   2973: 'Carrier 46 Power unit: Line phase failure in main circuit', class No Acknowledgement, trigger "DB302_HMI_Faults_Carrier46_Faults_1" bit 12
   2974: 'Carrier 46 Power unit: Phase failure motor cable', class No Acknowledgement, trigger "DB302_HMI_Faults_Carrier46_Faults_1" bit 13
   2975: 'Carrier 46 Power unit: Ground fault', class No Acknowledgement, trigger "DB302_HMI_Faults_Carrier46_Faults_1" bit 14
   2976: 'Spare_Fault_2976', class No Acknowledgement, trigger "DB302_HMI_Faults_Carrier46_Faults_1" bit 15
   2977: 'Carrier 46 Motion Off Fault', class No Acknowledgement, trigger "DB302_HMI_Faults_Carrier46_Faults_2" bit 0
   2978: 'Carrier 46 Motion On Fault', class No Acknowledgement, trigger "DB302_HMI_Faults_Carrier46_Faults_2" bit 1
   2979: 'Carrier 46 Spacing Fault', class No Acknowledgement, trigger "DB302_HMI_Faults_Carrier46_Faults_2" bit 2
   2980: 'Carrier 46 Duplicate Carrier Number Fault', class No Acknowledgement, trigger "DB302_HMI_Faults_Carrier46_Faults_2" bit 3
   2981: 'Spare_Fault_2981', class No Acknowledgement, trigger "DB302_HMI_Faults_Carrier46_Faults_2" bit 4
   2982: 'Spare_Fault_2982', class No Acknowledgement, trigger "DB302_HMI_Faults_Carrier46_Faults_2" bit 5
   2983: 'Spare_Fault_2983', class No Acknowledgement, trigger "DB302_HMI_Faults_Carrier46_Faults_2" bit 6
   2984: 'Spare_Fault_2984', class No Acknowledgement, trigger "DB302_HMI_Faults_Carrier46_Faults_2" bit 7
   2985: 'Spare_Fault_2985', class No Acknowledgement, trigger "DB302_HMI_Faults_Carrier46_Faults_2" bit 8
   2986: 'Spare_Fault_2986', class No Acknowledgement, trigger "DB302_HMI_Faults_Carrier46_Faults_2" bit 9
   2987: 'Spare_Fault_2987', class No Acknowledgement, trigger "DB302_HMI_Faults_Carrier46_Faults_2" bit 10
   2988: 'Spare_Fault_2988', class No Acknowledgement, trigger "DB302_HMI_Faults_Carrier46_Faults_2" bit 11
   2989: 'Spare_Fault_2989', class No Acknowledgement, trigger "DB302_HMI_Faults_Carrier46_Faults_2" bit 12
   2990: 'Spare_Fault_2990', class No Acknowledgement, trigger "DB302_HMI_Faults_Carrier46_Faults_2" bit 13
   2991: 'Spare_Fault_2991', class No Acknowledgement, trigger "DB302_HMI_Faults_Carrier46_Faults_2" bit 14
   2992: 'Spare_Fault_2992', class No Acknowledgement, trigger "DB302_HMI_Faults_Carrier46_Faults_2" bit 15
   2993: 'Spare_Fault_2993', class No Acknowledgement, trigger "DB302_HMI_Faults_Carrier46_Faults_3" bit 0
   2994: 'Spare_Fault_2994', class No Acknowledgement, trigger "DB302_HMI_Faults_Carrier46_Faults_3" bit 1
   2995: 'Spare_Fault_2995', class No Acknowledgement, trigger "DB302_HMI_Faults_Carrier46_Faults_3" bit 2
   2996: 'Spare_Fault_2996', class No Acknowledgement, trigger "DB302_HMI_Faults_Carrier46_Faults_3" bit 3
   2997: 'Spare_Fault_2997', class No Acknowledgement, trigger "DB302_HMI_Faults_Carrier46_Faults_3" bit 4
   2998: 'Spare_Fault_2998', class No Acknowledgement, trigger "DB302_HMI_Faults_Carrier46_Faults_3" bit 5
   2999: 'Spare_Fault_2999', class No Acknowledgement, trigger "DB302_HMI_Faults_Carrier46_Faults_3" bit 6
   3000: 'Spare_Fault_3000', class No Acknowledgement, trigger "DB302_HMI_Faults_Carrier46_Faults_3" bit 7
   3001: 'Spare_Fault_3001', class No Acknowledgement, trigger "DB302_HMI_Faults_Carrier46_Faults_3" bit 8
   3002: 'Spare_Fault_3002', class No Acknowledgement, trigger "DB302_HMI_Faults_Carrier46_Faults_3" bit 9
   3003: 'Spare_Fault_3003', class No Acknowledgement, trigger "DB302_HMI_Faults_Carrier46_Faults_3" bit 10
   3004: 'Spare_Fault_3004', class No Acknowledgement, trigger "DB302_HMI_Faults_Carrier46_Faults_3" bit 11
   3005: 'Spare_Fault_3005', class No Acknowledgement, trigger "DB302_HMI_Faults_Carrier46_Faults_3" bit 12
   3006: 'Spare_Fault_3006', class No Acknowledgement, trigger "DB302_HMI_Faults_Carrier46_Faults_3" bit 13
   3007: 'Spare_Fault_3007', class No Acknowledgement, trigger "DB302_HMI_Faults_Carrier46_Faults_3" bit 14
   3008: 'Spare_Fault_3008', class No Acknowledgement, trigger "DB302_HMI_Faults_Carrier46_Faults_3" bit 15
   3009: 'Carrier 47 Disconnect Open Power Fault DI11.0', class No Acknowledgement, trigger "DB302_HMI_Faults_Carrier47_Faults_0" bit 0
   3010: 'Carrier 47 Drive Profinet Comm Fault', class No Acknowledgement, trigger "DB302_HMI_Faults_Carrier47_Faults_0" bit 1
   3011: 'Carrier 47 Production Stop Not Reset', class No Acknowledgement, trigger "DB302_HMI_Faults_Carrier47_Faults_0" bit 2
   3012: 'Carrier 47 CB02122 Tripped', class No Acknowledgement, trigger "DB302_HMI_Faults_Carrier47_Faults_0" bit 3
   3013: 'Carrier 47 CB02123 Tripped', class No Acknowledgement, trigger "DB302_HMI_Faults_Carrier47_Faults_0" bit 4
   3014: 'Carrier 47 AUX1 CB Tripped', class No Acknowledgement, trigger "DB302_HMI_Faults_Carrier47_Faults_0" bit 5
   3015: 'Carrier 47 AUX2 CB Tripped', class No Acknowledgement, trigger "DB302_HMI_Faults_Carrier47_Faults_0" bit 6
   3016: 'Carrier 47 PLC Not Communicating', class No Acknowledgement, trigger "DB302_HMI_Faults_Carrier47_Faults_0" bit 7
   3017: 'Carrier 47 Safe Input Card Fault', class No Acknowledgement, trigger "DB302_HMI_Faults_Carrier47_Faults_0" bit 8
   3018: 'Carrier 47 Safe Output Card Fault', class No Acknowledgement, trigger "DB302_HMI_Faults_Carrier47_Faults_0" bit 9
   3019: 'Carrier 47 Standard Input Card Fault', class No Acknowledgement, trigger "DB302_HMI_Faults_Carrier47_Faults_0" bit 10
   3020: 'Carrier 47 Standard Output Card Fault', class No Acknowledgement, trigger "DB302_HMI_Faults_Carrier47_Faults_0" bit 11
   3021: 'Carrier 47 Encoder Position Fault', class No Acknowledgement, trigger "DB302_HMI_Faults_Carrier47_Faults_0" bit 12
   3022: 'Carrier 47 Encoder Internal Error', class No Acknowledgement, trigger "DB302_HMI_Faults_Carrier47_Faults_0" bit 13
   3023: 'Carrier 47 Encoder Comm Fault', class No Acknowledgement, trigger "DB302_HMI_Faults_Carrier47_Faults_0" bit 14
   3024: 'Carrier 47 HMI Comm Fault', class No Acknowledgement, trigger "DB302_HMI_Faults_Carrier47_Faults_0" bit 15
   3025: 'Carrier 47 Crash Detection Fault', class No Acknowledgement, trigger "DB302_HMI_Faults_Carrier47_Faults_1" bit 0
   3026: 'Carrier 47 Carrier Number Invalid', class No Acknowledgement, trigger "DB302_HMI_Faults_Carrier47_Faults_1" bit 1
   3027: 'Carrier 47 Drive: PROFINET configuration error', class No Acknowledgement, trigger "DB302_HMI_Faults_Carrier47_Faults_1" bit 2
   3028: 'Carrier 47 Drive: Error internal communications', class No Acknowledgement, trigger "DB302_HMI_Faults_Carrier47_Faults_1" bit 3
   3029: 'Carrier 47 Drive: Motor overtemperature', class No Acknowledgement, trigger "DB302_HMI_Faults_Carrier47_Faults_1" bit 4
   3030: 'Carrier 47 Drive: Motor overcurrent', class No Acknowledgement, trigger "DB302_HMI_Faults_Carrier47_Faults_1" bit 5
   3031: 'Carrier 47 Drive: Infeed or power unit not ready', class No Acknowledgement, trigger "DB302_HMI_Faults_Carrier47_Faults_1" bit 6
   3032: 'Carrier 47 Drive: Short-circuit/ground fault detected', class No Acknowledgement, trigger "DB302_HMI_Faults_Carrier47_Faults_1" bit 7
   3033: 'Carrier 47 Drive: PROFINET Setpoint timeout', class No Acknowledgement, trigger "DB302_HMI_Faults_Carrier47_Faults_1" bit 8
   3034: 'Carrier 47 Power unit: Overcurrent', class No Acknowledgement, trigger "DB302_HMI_Faults_Carrier47_Faults_1" bit 9
   3035: 'Carrier 47 Power unit: DC link voltage overvoltage', class No Acknowledgement, trigger "DB302_HMI_Faults_Carrier47_Faults_1" bit 10
   3036: 'Carrier 47 Power unit: DC link voltage undervoltage', class No Acknowledgement, trigger "DB302_HMI_Faults_Carrier47_Faults_1" bit 11
   3037: 'Carrier 47 Power unit: Line phase failure in main circuit', class No Acknowledgement, trigger "DB302_HMI_Faults_Carrier47_Faults_1" bit 12
   3038: 'Carrier 47 Power unit: Phase failure motor cable', class No Acknowledgement, trigger "DB302_HMI_Faults_Carrier47_Faults_1" bit 13
   3039: 'Carrier 47 Power unit: Ground fault', class No Acknowledgement, trigger "DB302_HMI_Faults_Carrier47_Faults_1" bit 14
   3040: 'Spare_Fault_3040', class No Acknowledgement, trigger "DB302_HMI_Faults_Carrier47_Faults_1" bit 15
   3041: 'Carrier 47 Motion Off Fault', class No Acknowledgement, trigger "DB302_HMI_Faults_Carrier47_Faults_2" bit 0
   3042: 'Carrier 47 Motion On Fault', class No Acknowledgement, trigger "DB302_HMI_Faults_Carrier47_Faults_2" bit 1
   3043: 'Carrier 47 Spacing Fault', class No Acknowledgement, trigger "DB302_HMI_Faults_Carrier47_Faults_2" bit 2
   3044: 'Carrier 47 Duplicate Carrier Number Fault', class No Acknowledgement, trigger "DB302_HMI_Faults_Carrier47_Faults_2" bit 3
   3045: 'Spare_Fault_3045', class No Acknowledgement, trigger "DB302_HMI_Faults_Carrier47_Faults_2" bit 4
   3046: 'Spare_Fault_3046', class No Acknowledgement, trigger "DB302_HMI_Faults_Carrier47_Faults_2" bit 5
   3047: 'Spare_Fault_3047', class No Acknowledgement, trigger "DB302_HMI_Faults_Carrier47_Faults_2" bit 6
   3048: 'Spare_Fault_3048', class No Acknowledgement, trigger "DB302_HMI_Faults_Carrier47_Faults_2" bit 7
   3049: 'Spare_Fault_3049', class No Acknowledgement, trigger "DB302_HMI_Faults_Carrier47_Faults_2" bit 8
   3050: 'Spare_Fault_3050', class No Acknowledgement, trigger "DB302_HMI_Faults_Carrier47_Faults_2" bit 9
   3051: 'Spare_Fault_3051', class No Acknowledgement, trigger "DB302_HMI_Faults_Carrier47_Faults_2" bit 10
   3052: 'Spare_Fault_3052', class No Acknowledgement, trigger "DB302_HMI_Faults_Carrier47_Faults_2" bit 11
   3053: 'Spare_Fault_3053', class No Acknowledgement, trigger "DB302_HMI_Faults_Carrier47_Faults_2" bit 12
   3054: 'Spare_Fault_3054', class No Acknowledgement, trigger "DB302_HMI_Faults_Carrier47_Faults_2" bit 13
   3055: 'Spare_Fault_3055', class No Acknowledgement, trigger "DB302_HMI_Faults_Carrier47_Faults_2" bit 14
   3056: 'Spare_Fault_3056', class No Acknowledgement, trigger "DB302_HMI_Faults_Carrier47_Faults_2" bit 15
   3057: 'Spare_Fault_3057', class No Acknowledgement, trigger "DB302_HMI_Faults_Carrier47_Faults_3" bit 0
   3058: 'Spare_Fault_3058', class No Acknowledgement, trigger "DB302_HMI_Faults_Carrier47_Faults_3" bit 1
   3059: 'Spare_Fault_3059', class No Acknowledgement, trigger "DB302_HMI_Faults_Carrier47_Faults_3" bit 2
   3060: 'Spare_Fault_3060', class No Acknowledgement, trigger "DB302_HMI_Faults_Carrier47_Faults_3" bit 3
   3061: 'Spare_Fault_3061', class No Acknowledgement, trigger "DB302_HMI_Faults_Carrier47_Faults_3" bit 4
   3062: 'Spare_Fault_3062', class No Acknowledgement, trigger "DB302_HMI_Faults_Carrier47_Faults_3" bit 5
   3063: 'Spare_Fault_3063', class No Acknowledgement, trigger "DB302_HMI_Faults_Carrier47_Faults_3" bit 6
   3064: 'Spare_Fault_3064', class No Acknowledgement, trigger "DB302_HMI_Faults_Carrier47_Faults_3" bit 7
   3065: 'Spare_Fault_3065', class No Acknowledgement, trigger "DB302_HMI_Faults_Carrier47_Faults_3" bit 8
   3066: 'Spare_Fault_3066', class No Acknowledgement, trigger "DB302_HMI_Faults_Carrier47_Faults_3" bit 9
   3067: 'Spare_Fault_3067', class No Acknowledgement, trigger "DB302_HMI_Faults_Carrier47_Faults_3" bit 10
   3068: 'Spare_Fault_3068', class No Acknowledgement, trigger "DB302_HMI_Faults_Carrier47_Faults_3" bit 11
   3069: 'Spare_Fault_3069', class No Acknowledgement, trigger "DB302_HMI_Faults_Carrier47_Faults_3" bit 12
   3070: 'Spare_Fault_3070', class No Acknowledgement, trigger "DB302_HMI_Faults_Carrier47_Faults_3" bit 13
   3071: 'Spare_Fault_3071', class No Acknowledgement, trigger "DB302_HMI_Faults_Carrier47_Faults_3" bit 14
   3072: 'Spare_Fault_3072', class No Acknowledgement, trigger "DB302_HMI_Faults_Carrier47_Faults_3" bit 15
   3073: 'Carrier 48 Disconnect Open Power Fault DI11.0', class No Acknowledgement, trigger "DB302_HMI_Faults_Carrier48_Faults_0" bit 0
   3074: 'Carrier 48 Drive Profinet Comm Fault', class No Acknowledgement, trigger "DB302_HMI_Faults_Carrier48_Faults_0" bit 1
   3075: 'Carrier 48 Production Stop Not Reset', class No Acknowledgement, trigger "DB302_HMI_Faults_Carrier48_Faults_0" bit 2
   3076: 'Carrier 48 CB02122 Tripped', class No Acknowledgement, trigger "DB302_HMI_Faults_Carrier48_Faults_0" bit 3
   3077: 'Carrier 48 CB02123 Tripped', class No Acknowledgement, trigger "DB302_HMI_Faults_Carrier48_Faults_0" bit 4
   3078: 'Carrier 48 AUX1 CB Tripped', class No Acknowledgement, trigger "DB302_HMI_Faults_Carrier48_Faults_0" bit 5
   3079: 'Carrier 48 AUX2 CB Tripped', class No Acknowledgement, trigger "DB302_HMI_Faults_Carrier48_Faults_0" bit 6
   3080: 'Carrier 48 PLC Not Communicating', class No Acknowledgement, trigger "DB302_HMI_Faults_Carrier48_Faults_0" bit 7
   3081: 'Carrier 48 Safe Input Card Fault', class No Acknowledgement, trigger "DB302_HMI_Faults_Carrier48_Faults_0" bit 8
   3082: 'Carrier 48 Safe Output Card Fault', class No Acknowledgement, trigger "DB302_HMI_Faults_Carrier48_Faults_0" bit 9
   3083: 'Carrier 48 Standard Input Card Fault', class No Acknowledgement, trigger "DB302_HMI_Faults_Carrier48_Faults_0" bit 10
   3084: 'Carrier 48 Standard Output Card Fault', class No Acknowledgement, trigger "DB302_HMI_Faults_Carrier48_Faults_0" bit 11
   3085: 'Carrier 48 Encoder Position Fault', class No Acknowledgement, trigger "DB302_HMI_Faults_Carrier48_Faults_0" bit 12
   3086: 'Carrier 48 Encoder Internal Error', class No Acknowledgement, trigger "DB302_HMI_Faults_Carrier48_Faults_0" bit 13
   3087: 'Carrier 48 Encoder Comm Fault', class No Acknowledgement, trigger "DB302_HMI_Faults_Carrier48_Faults_0" bit 14
   3088: 'Carrier 48 HMI Comm Fault', class No Acknowledgement, trigger "DB302_HMI_Faults_Carrier48_Faults_0" bit 15
   3089: 'Carrier 48 Crash Detection Fault', class No Acknowledgement, trigger "DB302_HMI_Faults_Carrier48_Faults_1" bit 0
   3090: 'Carrier 48 Carrier Number Invalid', class No Acknowledgement, trigger "DB302_HMI_Faults_Carrier48_Faults_1" bit 1
   3091: 'Carrier 48 Drive: PROFINET configuration error', class No Acknowledgement, trigger "DB302_HMI_Faults_Carrier48_Faults_1" bit 2
   3092: 'Carrier 48 Drive: Error internal communications', class No Acknowledgement, trigger "DB302_HMI_Faults_Carrier48_Faults_1" bit 3
   3093: 'Carrier 48 Drive: Motor overtemperature', class No Acknowledgement, trigger "DB302_HMI_Faults_Carrier48_Faults_1" bit 4
   3094: 'Carrier 48 Drive: Motor overcurrent', class No Acknowledgement, trigger "DB302_HMI_Faults_Carrier48_Faults_1" bit 5
   3095: 'Carrier 48 Drive: Infeed or power unit not ready', class No Acknowledgement, trigger "DB302_HMI_Faults_Carrier48_Faults_1" bit 6
   3096: 'Carrier 48 Drive: Short-circuit/ground fault detected', class No Acknowledgement, trigger "DB302_HMI_Faults_Carrier48_Faults_1" bit 7
   3097: 'Carrier 48 Drive: PROFINET Setpoint timeout', class No Acknowledgement, trigger "DB302_HMI_Faults_Carrier48_Faults_1" bit 8
   3098: 'Carrier 48 Power unit: Overcurrent', class No Acknowledgement, trigger "DB302_HMI_Faults_Carrier48_Faults_1" bit 9
   3099: 'Carrier 48 Power unit: DC link voltage overvoltage', class No Acknowledgement, trigger "DB302_HMI_Faults_Carrier48_Faults_1" bit 10
   3100: 'Carrier 48 Power unit: DC link voltage undervoltage', class No Acknowledgement, trigger "DB302_HMI_Faults_Carrier48_Faults_1" bit 11
   3101: 'Carrier 48 Power unit: Line phase failure in main circuit', class No Acknowledgement, trigger "DB302_HMI_Faults_Carrier48_Faults_1" bit 12
   3102: 'Carrier 48 Power unit: Phase failure motor cable', class No Acknowledgement, trigger "DB302_HMI_Faults_Carrier48_Faults_1" bit 13
   3103: 'Carrier 48 Power unit: Ground fault', class No Acknowledgement, trigger "DB302_HMI_Faults_Carrier48_Faults_1" bit 14
   3104: 'Spare_Fault_3104', class No Acknowledgement, trigger "DB302_HMI_Faults_Carrier48_Faults_1" bit 15
   3105: 'Carrier 48 Motion Off Fault', class No Acknowledgement, trigger "DB302_HMI_Faults_Carrier48_Faults_2" bit 0
   3106: 'Carrier 48 Motion On Fault', class No Acknowledgement, trigger "DB302_HMI_Faults_Carrier48_Faults_2" bit 1
   3107: 'Carrier 48 Spacing Fault', class No Acknowledgement, trigger "DB302_HMI_Faults_Carrier48_Faults_2" bit 2
   3108: 'Carrier 48 Duplicate Carrier Number Fault', class No Acknowledgement, trigger "DB302_HMI_Faults_Carrier48_Faults_2" bit 3
   3109: 'Spare_Fault_3109', class No Acknowledgement, trigger "DB302_HMI_Faults_Carrier48_Faults_2" bit 4
   3110: 'Spare_Fault_3110', class No Acknowledgement, trigger "DB302_HMI_Faults_Carrier48_Faults_2" bit 5
   3111: 'Spare_Fault_3111', class No Acknowledgement, trigger "DB302_HMI_Faults_Carrier48_Faults_2" bit 6
   3112: 'Spare_Fault_3112', class No Acknowledgement, trigger "DB302_HMI_Faults_Carrier48_Faults_2" bit 7
   3113: 'Spare_Fault_3113', class No Acknowledgement, trigger "DB302_HMI_Faults_Carrier48_Faults_2" bit 8
   3114: 'Spare_Fault_3114', class No Acknowledgement, trigger "DB302_HMI_Faults_Carrier48_Faults_2" bit 9
   3115: 'Spare_Fault_3115', class No Acknowledgement, trigger "DB302_HMI_Faults_Carrier48_Faults_2" bit 10
   3116: 'Spare_Fault_3116', class No Acknowledgement, trigger "DB302_HMI_Faults_Carrier48_Faults_2" bit 11
   3117: 'Spare_Fault_3117', class No Acknowledgement, trigger "DB302_HMI_Faults_Carrier48_Faults_2" bit 12
   3118: 'Spare_Fault_3118', class No Acknowledgement, trigger "DB302_HMI_Faults_Carrier48_Faults_2" bit 13
   3119: 'Spare_Fault_3119', class No Acknowledgement, trigger "DB302_HMI_Faults_Carrier48_Faults_2" bit 14
   3120: 'Spare_Fault_3120', class No Acknowledgement, trigger "DB302_HMI_Faults_Carrier48_Faults_2" bit 15
   3121: 'Spare_Fault_3121', class No Acknowledgement, trigger "DB302_HMI_Faults_Carrier48_Faults_3" bit 0
   3122: 'Spare_Fault_3122', class No Acknowledgement, trigger "DB302_HMI_Faults_Carrier48_Faults_3" bit 1
   3123: 'Spare_Fault_3123', class No Acknowledgement, trigger "DB302_HMI_Faults_Carrier48_Faults_3" bit 2
   3124: 'Spare_Fault_3124', class No Acknowledgement, trigger "DB302_HMI_Faults_Carrier48_Faults_3" bit 3
   3125: 'Spare_Fault_3125', class No Acknowledgement, trigger "DB302_HMI_Faults_Carrier48_Faults_3" bit 4
   3126: 'Spare_Fault_3126', class No Acknowledgement, trigger "DB302_HMI_Faults_Carrier48_Faults_3" bit 5
   3127: 'Spare_Fault_3127', class No Acknowledgement, trigger "DB302_HMI_Faults_Carrier48_Faults_3" bit 6
   3128: 'Spare_Fault_3128', class No Acknowledgement, trigger "DB302_HMI_Faults_Carrier48_Faults_3" bit 7
   3129: 'Spare_Fault_3129', class No Acknowledgement, trigger "DB302_HMI_Faults_Carrier48_Faults_3" bit 8
   3130: 'Spare_Fault_3130', class No Acknowledgement, trigger "DB302_HMI_Faults_Carrier48_Faults_3" bit 9
   3131: 'Spare_Fault_3131', class No Acknowledgement, trigger "DB302_HMI_Faults_Carrier48_Faults_3" bit 10
   3132: 'Spare_Fault_3132', class No Acknowledgement, trigger "DB302_HMI_Faults_Carrier48_Faults_3" bit 11
   3133: 'Spare_Fault_3133', class No Acknowledgement, trigger "DB302_HMI_Faults_Carrier48_Faults_3" bit 12
   3134: 'Spare_Fault_3134', class No Acknowledgement, trigger "DB302_HMI_Faults_Carrier48_Faults_3" bit 13
   3135: 'Spare_Fault_3135', class No Acknowledgement, trigger "DB302_HMI_Faults_Carrier48_Faults_3" bit 14
   3136: 'Spare_Fault_3136', class No Acknowledgement, trigger "DB302_HMI_Faults_Carrier48_Faults_3" bit 15
   3137: 'Carrier 49 Disconnect Open Power Fault DI11.0', class No Acknowledgement, trigger "DB302_HMI_Faults_Carrier49_Faults_0" bit 0
   3138: 'Carrier 49 Drive Profinet Comm Fault', class No Acknowledgement, trigger "DB302_HMI_Faults_Carrier49_Faults_0" bit 1
   3139: 'Carrier 49 Production Stop Not Reset', class No Acknowledgement, trigger "DB302_HMI_Faults_Carrier49_Faults_0" bit 2
   3140: 'Carrier 49 CB02122 Tripped', class No Acknowledgement, trigger "DB302_HMI_Faults_Carrier49_Faults_0" bit 3
   3141: 'Carrier 49 CB02123 Tripped', class No Acknowledgement, trigger "DB302_HMI_Faults_Carrier49_Faults_0" bit 4
   3142: 'Carrier 49 AUX1 CB Tripped', class No Acknowledgement, trigger "DB302_HMI_Faults_Carrier49_Faults_0" bit 5
   3143: 'Carrier 49 AUX2 CB Tripped', class No Acknowledgement, trigger "DB302_HMI_Faults_Carrier49_Faults_0" bit 6
   3144: 'Carrier 49 PLC Not Communicating', class No Acknowledgement, trigger "DB302_HMI_Faults_Carrier49_Faults_0" bit 7
   3145: 'Carrier 49 Safe Input Card Fault', class No Acknowledgement, trigger "DB302_HMI_Faults_Carrier49_Faults_0" bit 8
   3146: 'Carrier 49 Safe Output Card Fault', class No Acknowledgement, trigger "DB302_HMI_Faults_Carrier49_Faults_0" bit 9
   3147: 'Carrier 49 Standard Input Card Fault', class No Acknowledgement, trigger "DB302_HMI_Faults_Carrier49_Faults_0" bit 10
   3148: 'Carrier 49 Standard Output Card Fault', class No Acknowledgement, trigger "DB302_HMI_Faults_Carrier49_Faults_0" bit 11
   3149: 'Carrier 49 Encoder Position Fault', class No Acknowledgement, trigger "DB302_HMI_Faults_Carrier49_Faults_0" bit 12
   3150: 'Carrier 49 Encoder Internal Error', class No Acknowledgement, trigger "DB302_HMI_Faults_Carrier49_Faults_0" bit 13
   3151: 'Carrier 49 Encoder Comm Fault', class No Acknowledgement, trigger "DB302_HMI_Faults_Carrier49_Faults_0" bit 14
   3152: 'Carrier 49 HMI Comm Fault', class No Acknowledgement, trigger "DB302_HMI_Faults_Carrier49_Faults_0" bit 15
   3153: 'Carrier 49 Crash Detection Fault', class No Acknowledgement, trigger "DB302_HMI_Faults_Carrier49_Faults_1" bit 0
   3154: 'Carrier 49 Carrier Number Invalid', class No Acknowledgement, trigger "DB302_HMI_Faults_Carrier49_Faults_1" bit 1
   3155: 'Carrier 49 Drive: PROFINET configuration error', class No Acknowledgement, trigger "DB302_HMI_Faults_Carrier49_Faults_1" bit 2
   3156: 'Carrier 49 Drive: Error internal communications', class No Acknowledgement, trigger "DB302_HMI_Faults_Carrier49_Faults_1" bit 3
   3157: 'Carrier 49 Drive: Motor overtemperature', class No Acknowledgement, trigger "DB302_HMI_Faults_Carrier49_Faults_1" bit 4
   3158: 'Carrier 49 Drive: Motor overcurrent', class No Acknowledgement, trigger "DB302_HMI_Faults_Carrier49_Faults_1" bit 5
   3159: 'Carrier 49 Drive: Infeed or power unit not ready', class No Acknowledgement, trigger "DB302_HMI_Faults_Carrier49_Faults_1" bit 6
   3160: 'Carrier 49 Drive: Short-circuit/ground fault detected', class No Acknowledgement, trigger "DB302_HMI_Faults_Carrier49_Faults_1" bit 7
   3161: 'Carrier 49 Drive: PROFINET Setpoint timeout', class No Acknowledgement, trigger "DB302_HMI_Faults_Carrier49_Faults_1" bit 8
   3162: 'Carrier 49 Power unit: Overcurrent', class No Acknowledgement, trigger "DB302_HMI_Faults_Carrier49_Faults_1" bit 9
   3163: 'Carrier 49 Power unit: DC link voltage overvoltage', class No Acknowledgement, trigger "DB302_HMI_Faults_Carrier49_Faults_1" bit 10
   3164: 'Carrier 49 Power unit: DC link voltage undervoltage', class No Acknowledgement, trigger "DB302_HMI_Faults_Carrier49_Faults_1" bit 11
   3165: 'Carrier 49 Power unit: Line phase failure in main circuit', class No Acknowledgement, trigger "DB302_HMI_Faults_Carrier49_Faults_1" bit 12
   3166: 'Carrier 49 Power unit: Phase failure motor cable', class No Acknowledgement, trigger "DB302_HMI_Faults_Carrier49_Faults_1" bit 13
   3167: 'Carrier 49 Power unit: Ground fault', class No Acknowledgement, trigger "DB302_HMI_Faults_Carrier49_Faults_1" bit 14
   3168: 'Spare_Fault_3168', class No Acknowledgement, trigger "DB302_HMI_Faults_Carrier49_Faults_1" bit 15
   3169: 'Carrier 49 Motion Off Fault', class No Acknowledgement, trigger "DB302_HMI_Faults_Carrier49_Faults_2" bit 0
   3170: 'Carrier 49 Motion On Fault', class No Acknowledgement, trigger "DB302_HMI_Faults_Carrier49_Faults_2" bit 1
   3171: 'Carrier 49 Spacing Fault', class No Acknowledgement, trigger "DB302_HMI_Faults_Carrier49_Faults_2" bit 2
   3172: 'Carrier 49 Duplicate Carrier Number Fault', class No Acknowledgement, trigger "DB302_HMI_Faults_Carrier49_Faults_2" bit 3
   3173: 'Spare_Fault_3173', class No Acknowledgement, trigger "DB302_HMI_Faults_Carrier49_Faults_2" bit 4
   3174: 'Spare_Fault_3174', class No Acknowledgement, trigger "DB302_HMI_Faults_Carrier49_Faults_2" bit 5
   3175: 'Spare_Fault_3175', class No Acknowledgement, trigger "DB302_HMI_Faults_Carrier49_Faults_2" bit 6
   3176: 'Spare_Fault_3176', class No Acknowledgement, trigger "DB302_HMI_Faults_Carrier49_Faults_2" bit 7
   3177: 'Spare_Fault_3177', class No Acknowledgement, trigger "DB302_HMI_Faults_Carrier49_Faults_2" bit 8
   3178: 'Spare_Fault_3178', class No Acknowledgement, trigger "DB302_HMI_Faults_Carrier49_Faults_2" bit 9
   3179: 'Spare_Fault_3179', class No Acknowledgement, trigger "DB302_HMI_Faults_Carrier49_Faults_2" bit 10
   3180: 'Spare_Fault_3180', class No Acknowledgement, trigger "DB302_HMI_Faults_Carrier49_Faults_2" bit 11
   3181: 'Spare_Fault_3181', class No Acknowledgement, trigger "DB302_HMI_Faults_Carrier49_Faults_2" bit 12
   3182: 'Spare_Fault_3182', class No Acknowledgement, trigger "DB302_HMI_Faults_Carrier49_Faults_2" bit 13
   3183: 'Spare_Fault_3183', class No Acknowledgement, trigger "DB302_HMI_Faults_Carrier49_Faults_2" bit 14
   3184: 'Spare_Fault_3184', class No Acknowledgement, trigger "DB302_HMI_Faults_Carrier49_Faults_2" bit 15
   3185: 'Spare_Fault_3185', class No Acknowledgement, trigger "DB302_HMI_Faults_Carrier49_Faults_3" bit 0
   3186: 'Spare_Fault_3186', class No Acknowledgement, trigger "DB302_HMI_Faults_Carrier49_Faults_3" bit 1
   3187: 'Spare_Fault_3187', class No Acknowledgement, trigger "DB302_HMI_Faults_Carrier49_Faults_3" bit 2
   3188: 'Spare_Fault_3188', class No Acknowledgement, trigger "DB302_HMI_Faults_Carrier49_Faults_3" bit 3
   3189: 'Spare_Fault_3189', class No Acknowledgement, trigger "DB302_HMI_Faults_Carrier49_Faults_3" bit 4
   3190: 'Spare_Fault_3190', class No Acknowledgement, trigger "DB302_HMI_Faults_Carrier49_Faults_3" bit 5
   3191: 'Spare_Fault_3191', class No Acknowledgement, trigger "DB302_HMI_Faults_Carrier49_Faults_3" bit 6
   3192: 'Spare_Fault_3192', class No Acknowledgement, trigger "DB302_HMI_Faults_Carrier49_Faults_3" bit 7
   3193: 'Spare_Fault_3193', class No Acknowledgement, trigger "DB302_HMI_Faults_Carrier49_Faults_3" bit 8
   3194: 'Spare_Fault_3194', class No Acknowledgement, trigger "DB302_HMI_Faults_Carrier49_Faults_3" bit 9
   3195: 'Spare_Fault_3195', class No Acknowledgement, trigger "DB302_HMI_Faults_Carrier49_Faults_3" bit 10
   3196: 'Spare_Fault_3196', class No Acknowledgement, trigger "DB302_HMI_Faults_Carrier49_Faults_3" bit 11
   3197: 'Spare_Fault_3197', class No Acknowledgement, trigger "DB302_HMI_Faults_Carrier49_Faults_3" bit 12
   3198: 'Spare_Fault_3198', class No Acknowledgement, trigger "DB302_HMI_Faults_Carrier49_Faults_3" bit 13
   3199: 'Spare_Fault_3199', class No Acknowledgement, trigger "DB302_HMI_Faults_Carrier49_Faults_3" bit 14
   3200: 'Spare_Fault_3200', class No Acknowledgement, trigger "DB302_HMI_Faults_Carrier49_Faults_3" bit 15
   3201: 'Carrier 50 Disconnect Open Power Fault DI11.0', class No Acknowledgement, trigger "DB302_HMI_Faults_Carrier50_Faults_0" bit 0
   3202: 'Carrier 50 Drive Profinet Comm Fault', class No Acknowledgement, trigger "DB302_HMI_Faults_Carrier50_Faults_0" bit 1
   3203: 'Carrier 50 Production Stop Not Reset', class No Acknowledgement, trigger "DB302_HMI_Faults_Carrier50_Faults_0" bit 2
   3204: 'Carrier 50 CB02122 Tripped', class No Acknowledgement, trigger "DB302_HMI_Faults_Carrier50_Faults_0" bit 3
   3205: 'Carrier 50 CB02123 Tripped', class No Acknowledgement, trigger "DB302_HMI_Faults_Carrier50_Faults_0" bit 4
   3206: 'Carrier 50 AUX1 CB Tripped', class No Acknowledgement, trigger "DB302_HMI_Faults_Carrier50_Faults_0" bit 5
   3207: 'Carrier 50 AUX2 CB Tripped', class No Acknowledgement, trigger "DB302_HMI_Faults_Carrier50_Faults_0" bit 6
   3208: 'Carrier 50 PLC Not Communicating', class No Acknowledgement, trigger "DB302_HMI_Faults_Carrier50_Faults_0" bit 7
   3209: 'Carrier 50 Safe Input Card Fault', class No Acknowledgement, trigger "DB302_HMI_Faults_Carrier50_Faults_0" bit 8
   3210: 'Carrier 50 Safe Output Card Fault', class No Acknowledgement, trigger "DB302_HMI_Faults_Carrier50_Faults_0" bit 9
   3211: 'Carrier 50 Standard Input Card Fault', class No Acknowledgement, trigger "DB302_HMI_Faults_Carrier50_Faults_0" bit 10
   3212: 'Carrier 50 Standard Output Card Fault', class No Acknowledgement, trigger "DB302_HMI_Faults_Carrier50_Faults_0" bit 11
   3213: 'Carrier 50 Encoder Position Fault', class No Acknowledgement, trigger "DB302_HMI_Faults_Carrier50_Faults_0" bit 12
   3214: 'Carrier 50 Encoder Internal Error', class No Acknowledgement, trigger "DB302_HMI_Faults_Carrier50_Faults_0" bit 13
   3215: 'Carrier 50 Encoder Comm Fault', class No Acknowledgement, trigger "DB302_HMI_Faults_Carrier50_Faults_0" bit 14
   3216: 'Carrier 50 HMI Comm Fault', class No Acknowledgement, trigger "DB302_HMI_Faults_Carrier50_Faults_0" bit 15
   3217: 'Carrier 50 Crash Detection Fault', class No Acknowledgement, trigger "DB302_HMI_Faults_Carrier50_Faults_1" bit 0
   3218: 'Carrier 50 Carrier Number Invalid', class No Acknowledgement, trigger "DB302_HMI_Faults_Carrier50_Faults_1" bit 1
   3219: 'Carrier 50 Drive: PROFINET configuration error', class No Acknowledgement, trigger "DB302_HMI_Faults_Carrier50_Faults_1" bit 2
   3220: 'Carrier 50 Drive: Error internal communications', class No Acknowledgement, trigger "DB302_HMI_Faults_Carrier50_Faults_1" bit 3
   3221: 'Carrier 50 Drive: Motor overtemperature', class No Acknowledgement, trigger "DB302_HMI_Faults_Carrier50_Faults_1" bit 4
   3222: 'Carrier 50 Drive: Motor overcurrent', class No Acknowledgement, trigger "DB302_HMI_Faults_Carrier50_Faults_1" bit 5
   3223: 'Carrier 50 Drive: Infeed or power unit not ready', class No Acknowledgement, trigger "DB302_HMI_Faults_Carrier50_Faults_1" bit 6
   3224: 'Carrier 50 Drive: Short-circuit/ground fault detected', class No Acknowledgement, trigger "DB302_HMI_Faults_Carrier50_Faults_1" bit 7
   3225: 'Carrier 50 Drive: PROFINET Setpoint timeout', class No Acknowledgement, trigger "DB302_HMI_Faults_Carrier50_Faults_1" bit 8
   3226: 'Carrier 50 Power unit: Overcurrent', class No Acknowledgement, trigger "DB302_HMI_Faults_Carrier50_Faults_1" bit 9
   3227: 'Carrier 50 Power unit: DC link voltage overvoltage', class No Acknowledgement, trigger "DB302_HMI_Faults_Carrier50_Faults_1" bit 10
   3228: 'Carrier 50 Power unit: DC link voltage undervoltage', class No Acknowledgement, trigger "DB302_HMI_Faults_Carrier50_Faults_1" bit 11
   3229: 'Carrier 50 Power unit: Line phase failure in main circuit', class No Acknowledgement, trigger "DB302_HMI_Faults_Carrier50_Faults_1" bit 12
   3230: 'Carrier 50 Power unit: Phase failure motor cable', class No Acknowledgement, trigger "DB302_HMI_Faults_Carrier50_Faults_1" bit 13
   3231: 'Carrier 50 Power unit: Ground fault', class No Acknowledgement, trigger "DB302_HMI_Faults_Carrier50_Faults_1" bit 14
   3232: 'Spare_Fault_3232', class No Acknowledgement, trigger "DB302_HMI_Faults_Carrier50_Faults_1" bit 15
   3233: 'Carrier 50 Motion Off Fault', class No Acknowledgement, trigger "DB302_HMI_Faults_Carrier50_Faults_2" bit 0
   3234: 'Carrier 50 Motion On Fault', class No Acknowledgement, trigger "DB302_HMI_Faults_Carrier50_Faults_2" bit 1
   3235: 'Carrier 50 Spacing Fault', class No Acknowledgement, trigger "DB302_HMI_Faults_Carrier50_Faults_2" bit 2
   3236: 'Carrier 50 Duplicate Carrier Number Fault', class No Acknowledgement, trigger "DB302_HMI_Faults_Carrier50_Faults_2" bit 3
   3237: 'Spare_Fault_3237', class No Acknowledgement, trigger "DB302_HMI_Faults_Carrier50_Faults_2" bit 4
   3238: 'Spare_Fault_3238', class No Acknowledgement, trigger "DB302_HMI_Faults_Carrier50_Faults_2" bit 5
   3239: 'Spare_Fault_3239', class No Acknowledgement, trigger "DB302_HMI_Faults_Carrier50_Faults_2" bit 6
   3240: 'Spare_Fault_3240', class No Acknowledgement, trigger "DB302_HMI_Faults_Carrier50_Faults_2" bit 7
   3241: 'Spare_Fault_3241', class No Acknowledgement, trigger "DB302_HMI_Faults_Carrier50_Faults_2" bit 8
   3242: 'Spare_Fault_3242', class No Acknowledgement, trigger "DB302_HMI_Faults_Carrier50_Faults_2" bit 9
   3243: 'Spare_Fault_3243', class No Acknowledgement, trigger "DB302_HMI_Faults_Carrier50_Faults_2" bit 10
   3244: 'Spare_Fault_3244', class No Acknowledgement, trigger "DB302_HMI_Faults_Carrier50_Faults_2" bit 11
   3245: 'Spare_Fault_3245', class No Acknowledgement, trigger "DB302_HMI_Faults_Carrier50_Faults_2" bit 12
   3246: 'Spare_Fault_3246', class No Acknowledgement, trigger "DB302_HMI_Faults_Carrier50_Faults_2" bit 13
   3247: 'Spare_Fault_3247', class No Acknowledgement, trigger "DB302_HMI_Faults_Carrier50_Faults_2" bit 14
   3248: 'Spare_Fault_3248', class No Acknowledgement, trigger "DB302_HMI_Faults_Carrier50_Faults_2" bit 15
   3249: 'Spare_Fault_3249', class No Acknowledgement, trigger "DB302_HMI_Faults_Carrier50_Faults_3" bit 0
   3250: 'Spare_Fault_3250', class No Acknowledgement, trigger "DB302_HMI_Faults_Carrier50_Faults_3" bit 1
   3251: 'Spare_Fault_3251', class No Acknowledgement, trigger "DB302_HMI_Faults_Carrier50_Faults_3" bit 2
   3252: 'Spare_Fault_3252', class No Acknowledgement, trigger "DB302_HMI_Faults_Carrier50_Faults_3" bit 3
   3253: 'Spare_Fault_3253', class No Acknowledgement, trigger "DB302_HMI_Faults_Carrier50_Faults_3" bit 4
   3254: 'Spare_Fault_3254', class No Acknowledgement, trigger "DB302_HMI_Faults_Carrier50_Faults_3" bit 5
   3255: 'Spare_Fault_3255', class No Acknowledgement, trigger "DB302_HMI_Faults_Carrier50_Faults_3" bit 6
   3256: 'Spare_Fault_3256', class No Acknowledgement, trigger "DB302_HMI_Faults_Carrier50_Faults_3" bit 7
   3257: 'Spare_Fault_3257', class No Acknowledgement, trigger "DB302_HMI_Faults_Carrier50_Faults_3" bit 8
   3258: 'Spare_Fault_3258', class No Acknowledgement, trigger "DB302_HMI_Faults_Carrier50_Faults_3" bit 9
   3259: 'Spare_Fault_3259', class No Acknowledgement, trigger "DB302_HMI_Faults_Carrier50_Faults_3" bit 10
   3260: 'Spare_Fault_3260', class No Acknowledgement, trigger "DB302_HMI_Faults_Carrier50_Faults_3" bit 11
   3261: 'Spare_Fault_3261', class No Acknowledgement, trigger "DB302_HMI_Faults_Carrier50_Faults_3" bit 12
   3262: 'Spare_Fault_3262', class No Acknowledgement, trigger "DB302_HMI_Faults_Carrier50_Faults_3" bit 13
   3263: 'Spare_Fault_3263', class No Acknowledgement, trigger "DB302_HMI_Faults_Carrier50_Faults_3" bit 14
   3264: 'Spare_Fault_3264', class No Acknowledgement, trigger "DB302_HMI_Faults_Carrier50_Faults_3" bit 15
   3265: 'Carrier 51 Disconnect Open Power Fault DI11.0', class No Acknowledgement, trigger "DB302_HMI_Faults_Carrier51_Faults_0" bit 0
   3266: 'Carrier 51 Drive Profinet Comm Fault', class No Acknowledgement, trigger "DB302_HMI_Faults_Carrier51_Faults_0" bit 1
   3267: 'Carrier 51 Production Stop Not Reset', class No Acknowledgement, trigger "DB302_HMI_Faults_Carrier51_Faults_0" bit 2
   3268: 'Carrier 51 CB02122 Tripped', class No Acknowledgement, trigger "DB302_HMI_Faults_Carrier51_Faults_0" bit 3
   3269: 'Carrier 51 CB02123 Tripped', class No Acknowledgement, trigger "DB302_HMI_Faults_Carrier51_Faults_0" bit 4
   3270: 'Carrier 51 AUX1 CB Tripped', class No Acknowledgement, trigger "DB302_HMI_Faults_Carrier51_Faults_0" bit 5
   3271: 'Carrier 51 AUX2 CB Tripped', class No Acknowledgement, trigger "DB302_HMI_Faults_Carrier51_Faults_0" bit 6
   3272: 'Carrier 51 PLC Not Communicating', class No Acknowledgement, trigger "DB302_HMI_Faults_Carrier51_Faults_0" bit 7
   3273: 'Carrier 51 Safe Input Card Fault', class No Acknowledgement, trigger "DB302_HMI_Faults_Carrier51_Faults_0" bit 8
   3274: 'Carrier 51 Safe Output Card Fault', class No Acknowledgement, trigger "DB302_HMI_Faults_Carrier51_Faults_0" bit 9
   3275: 'Carrier 51 Standard Input Card Fault', class No Acknowledgement, trigger "DB302_HMI_Faults_Carrier51_Faults_0" bit 10
   3276: 'Carrier 51 Standard Output Card Fault', class No Acknowledgement, trigger "DB302_HMI_Faults_Carrier51_Faults_0" bit 11
   3277: 'Carrier 51 Encoder Position Fault', class No Acknowledgement, trigger "DB302_HMI_Faults_Carrier51_Faults_0" bit 12
   3278: 'Carrier 51 Encoder Internal Error', class No Acknowledgement, trigger "DB302_HMI_Faults_Carrier51_Faults_0" bit 13
   3279: 'Carrier 51 Encoder Comm Fault', class No Acknowledgement, trigger "DB302_HMI_Faults_Carrier51_Faults_0" bit 14
   3280: 'Carrier 51 HMI Comm Fault', class No Acknowledgement, trigger "DB302_HMI_Faults_Carrier51_Faults_0" bit 15
   3281: 'Carrier 51 Crash Detection Fault', class No Acknowledgement, trigger "DB302_HMI_Faults_Carrier51_Faults_1" bit 0
   3282: 'Carrier 51 Carrier Number Invalid', class No Acknowledgement, trigger "DB302_HMI_Faults_Carrier51_Faults_1" bit 1
   3283: 'Carrier 51 Drive: PROFINET configuration error', class No Acknowledgement, trigger "DB302_HMI_Faults_Carrier51_Faults_1" bit 2
   3284: 'Carrier 51 Drive: Error internal communications', class No Acknowledgement, trigger "DB302_HMI_Faults_Carrier51_Faults_1" bit 3
   3285: 'Carrier 51 Drive: Motor overtemperature', class No Acknowledgement, trigger "DB302_HMI_Faults_Carrier51_Faults_1" bit 4
   3286: 'Carrier 51 Drive: Motor overcurrent', class No Acknowledgement, trigger "DB302_HMI_Faults_Carrier51_Faults_1" bit 5
   3287: 'Carrier 51 Drive: Infeed or power unit not ready', class No Acknowledgement, trigger "DB302_HMI_Faults_Carrier51_Faults_1" bit 6
   3288: 'Carrier 51 Drive: Short-circuit/ground fault detected', class No Acknowledgement, trigger "DB302_HMI_Faults_Carrier51_Faults_1" bit 7
   3289: 'Carrier 51 Drive: PROFINET Setpoint timeout', class No Acknowledgement, trigger "DB302_HMI_Faults_Carrier51_Faults_1" bit 8
   3290: 'Carrier 51 Power unit: Overcurrent', class No Acknowledgement, trigger "DB302_HMI_Faults_Carrier51_Faults_1" bit 9
   3291: 'Carrier 51 Power unit: DC link voltage overvoltage', class No Acknowledgement, trigger "DB302_HMI_Faults_Carrier51_Faults_1" bit 10
   3292: 'Carrier 51 Power unit: DC link voltage undervoltage', class No Acknowledgement, trigger "DB302_HMI_Faults_Carrier51_Faults_1" bit 11
   3293: 'Carrier 51 Power unit: Line phase failure in main circuit', class No Acknowledgement, trigger "DB302_HMI_Faults_Carrier51_Faults_1" bit 12
   3294: 'Carrier 51 Power unit: Phase failure motor cable', class No Acknowledgement, trigger "DB302_HMI_Faults_Carrier51_Faults_1" bit 13
   3295: 'Carrier 51 Power unit: Ground fault', class No Acknowledgement, trigger "DB302_HMI_Faults_Carrier51_Faults_1" bit 14
   3296: 'Spare_Fault_3296', class No Acknowledgement, trigger "DB302_HMI_Faults_Carrier51_Faults_1" bit 15
   3297: 'Carrier 51 Motion Off Fault', class No Acknowledgement, trigger "DB302_HMI_Faults_Carrier51_Faults_2" bit 0
   3298: 'Carrier 51 Motion On Fault', class No Acknowledgement, trigger "DB302_HMI_Faults_Carrier51_Faults_2" bit 1
   3299: 'Carrier 51 Spacing Fault', class No Acknowledgement, trigger "DB302_HMI_Faults_Carrier51_Faults_2" bit 2
   3300: 'Carrier 51 Duplicate Carrier Number Fault', class No Acknowledgement, trigger "DB302_HMI_Faults_Carrier51_Faults_2" bit 3
   3301: 'Spare_Fault_3301', class No Acknowledgement, trigger "DB302_HMI_Faults_Carrier51_Faults_2" bit 4
   3302: 'Spare_Fault_3302', class No Acknowledgement, trigger "DB302_HMI_Faults_Carrier51_Faults_2" bit 5
   3303: 'Spare_Fault_3303', class No Acknowledgement, trigger "DB302_HMI_Faults_Carrier51_Faults_2" bit 6
   3304: 'Spare_Fault_3304', class No Acknowledgement, trigger "DB302_HMI_Faults_Carrier51_Faults_2" bit 7
   3305: 'Spare_Fault_3305', class No Acknowledgement, trigger "DB302_HMI_Faults_Carrier51_Faults_2" bit 8
   3306: 'Spare_Fault_3306', class No Acknowledgement, trigger "DB302_HMI_Faults_Carrier51_Faults_2" bit 9
   3307: 'Spare_Fault_3307', class No Acknowledgement, trigger "DB302_HMI_Faults_Carrier51_Faults_2" bit 10
   3308: 'Spare_Fault_3308', class No Acknowledgement, trigger "DB302_HMI_Faults_Carrier51_Faults_2" bit 11
   3309: 'Spare_Fault_3309', class No Acknowledgement, trigger "DB302_HMI_Faults_Carrier51_Faults_2" bit 12
   3310: 'Spare_Fault_3310', class No Acknowledgement, trigger "DB302_HMI_Faults_Carrier51_Faults_2" bit 13
   3311: 'Spare_Fault_3311', class No Acknowledgement, trigger "DB302_HMI_Faults_Carrier51_Faults_2" bit 14
   3312: 'Spare_Fault_3312', class No Acknowledgement, trigger "DB302_HMI_Faults_Carrier51_Faults_2" bit 15
   3313: 'Spare_Fault_3313', class No Acknowledgement, trigger "DB302_HMI_Faults_Carrier51_Faults_3" bit 0
   3314: 'Spare_Fault_3314', class No Acknowledgement, trigger "DB302_HMI_Faults_Carrier51_Faults_3" bit 1
   3315: 'Spare_Fault_3315', class No Acknowledgement, trigger "DB302_HMI_Faults_Carrier51_Faults_3" bit 2
   3316: 'Spare_Fault_3316', class No Acknowledgement, trigger "DB302_HMI_Faults_Carrier51_Faults_3" bit 3
   3317: 'Spare_Fault_3317', class No Acknowledgement, trigger "DB302_HMI_Faults_Carrier51_Faults_3" bit 4
   3318: 'Spare_Fault_3318', class No Acknowledgement, trigger "DB302_HMI_Faults_Carrier51_Faults_3" bit 5
   3319: 'Spare_Fault_3319', class No Acknowledgement, trigger "DB302_HMI_Faults_Carrier51_Faults_3" bit 6
   3320: 'Spare_Fault_3320', class No Acknowledgement, trigger "DB302_HMI_Faults_Carrier51_Faults_3" bit 7
   3321: 'Spare_Fault_3321', class No Acknowledgement, trigger "DB302_HMI_Faults_Carrier51_Faults_3" bit 8
   3322: 'Spare_Fault_3322', class No Acknowledgement, trigger "DB302_HMI_Faults_Carrier51_Faults_3" bit 9
   3323: 'Spare_Fault_3323', class No Acknowledgement, trigger "DB302_HMI_Faults_Carrier51_Faults_3" bit 10
   3324: 'Spare_Fault_3324', class No Acknowledgement, trigger "DB302_HMI_Faults_Carrier51_Faults_3" bit 11
   3325: 'Spare_Fault_3325', class No Acknowledgement, trigger "DB302_HMI_Faults_Carrier51_Faults_3" bit 12
   3326: 'Spare_Fault_3326', class No Acknowledgement, trigger "DB302_HMI_Faults_Carrier51_Faults_3" bit 13
   3327: 'Spare_Fault_3327', class No Acknowledgement, trigger "DB302_HMI_Faults_Carrier51_Faults_3" bit 14
   3328: 'Spare_Fault_3328', class No Acknowledgement, trigger "DB302_HMI_Faults_Carrier51_Faults_3" bit 15
   3329: 'Carrier 52 Disconnect Open Power Fault DI11.0', class No Acknowledgement, trigger "DB302_HMI_Faults_Carrier52_Faults_0" bit 0
   3330: 'Carrier 52 Drive Profinet Comm Fault', class No Acknowledgement, trigger "DB302_HMI_Faults_Carrier52_Faults_0" bit 1
   3331: 'Carrier 52 Production Stop Not Reset', class No Acknowledgement, trigger "DB302_HMI_Faults_Carrier52_Faults_0" bit 2
   3332: 'Carrier 52 CB02122 Tripped', class No Acknowledgement, trigger "DB302_HMI_Faults_Carrier52_Faults_0" bit 3
   3333: 'Carrier 52 CB02123 Tripped', class No Acknowledgement, trigger "DB302_HMI_Faults_Carrier52_Faults_0" bit 4
   3334: 'Carrier 52 AUX1 CB Tripped', class No Acknowledgement, trigger "DB302_HMI_Faults_Carrier52_Faults_0" bit 5
   3335: 'Carrier 52 AUX2 CB Tripped', class No Acknowledgement, trigger "DB302_HMI_Faults_Carrier52_Faults_0" bit 6
   3336: 'Carrier 52 PLC Not Communicating', class No Acknowledgement, trigger "DB302_HMI_Faults_Carrier52_Faults_0" bit 7
   3337: 'Carrier 52 Safe Input Card Fault', class No Acknowledgement, trigger "DB302_HMI_Faults_Carrier52_Faults_0" bit 8
   3338: 'Carrier 52 Safe Output Card Fault', class No Acknowledgement, trigger "DB302_HMI_Faults_Carrier52_Faults_0" bit 9
   3339: 'Carrier 52 Standard Input Card Fault', class No Acknowledgement, trigger "DB302_HMI_Faults_Carrier52_Faults_0" bit 10
   3340: 'Carrier 52 Standard Output Card Fault', class No Acknowledgement, trigger "DB302_HMI_Faults_Carrier52_Faults_0" bit 11
   3341: 'Carrier 52 Encoder Position Fault', class No Acknowledgement, trigger "DB302_HMI_Faults_Carrier52_Faults_0" bit 12
   3342: 'Carrier 52 Encoder Internal Error', class No Acknowledgement, trigger "DB302_HMI_Faults_Carrier52_Faults_0" bit 13
   3343: 'Carrier 52 Encoder Comm Fault', class No Acknowledgement, trigger "DB302_HMI_Faults_Carrier52_Faults_0" bit 14
   3344: 'Carrier 52 HMI Comm Fault', class No Acknowledgement, trigger "DB302_HMI_Faults_Carrier52_Faults_0" bit 15
   3345: 'Carrier 52 Crash Detection Fault', class No Acknowledgement, trigger "DB302_HMI_Faults_Carrier52_Faults_1" bit 0
   3346: 'Carrier 52 Carrier Number Invalid', class No Acknowledgement, trigger "DB302_HMI_Faults_Carrier52_Faults_1" bit 1
   3347: 'Carrier 52 Drive: PROFINET configuration error', class No Acknowledgement, trigger "DB302_HMI_Faults_Carrier52_Faults_1" bit 2
   3348: 'Carrier 52 Drive: Error internal communications', class No Acknowledgement, trigger "DB302_HMI_Faults_Carrier52_Faults_1" bit 3
   3349: 'Carrier 52 Drive: Motor overtemperature', class No Acknowledgement, trigger "DB302_HMI_Faults_Carrier52_Faults_1" bit 4
   3350: 'Carrier 52 Drive: Motor overcurrent', class No Acknowledgement, trigger "DB302_HMI_Faults_Carrier52_Faults_1" bit 5
   3351: 'Carrier 52 Drive: Infeed or power unit not ready', class No Acknowledgement, trigger "DB302_HMI_Faults_Carrier52_Faults_1" bit 6
   3352: 'Carrier 52 Drive: Short-circuit/ground fault detected', class No Acknowledgement, trigger "DB302_HMI_Faults_Carrier52_Faults_1" bit 7
   3353: 'Carrier 52 Drive: PROFINET Setpoint timeout', class No Acknowledgement, trigger "DB302_HMI_Faults_Carrier52_Faults_1" bit 8
   3354: 'Carrier 52 Power unit: Overcurrent', class No Acknowledgement, trigger "DB302_HMI_Faults_Carrier52_Faults_1" bit 9
   3355: 'Carrier 52 Power unit: DC link voltage overvoltage', class No Acknowledgement, trigger "DB302_HMI_Faults_Carrier52_Faults_1" bit 10
   3356: 'Carrier 52 Power unit: DC link voltage undervoltage', class No Acknowledgement, trigger "DB302_HMI_Faults_Carrier52_Faults_1" bit 11
   3357: 'Carrier 52 Power unit: Line phase failure in main circuit', class No Acknowledgement, trigger "DB302_HMI_Faults_Carrier52_Faults_1" bit 12
   3358: 'Carrier 52 Power unit: Phase failure motor cable', class No Acknowledgement, trigger "DB302_HMI_Faults_Carrier52_Faults_1" bit 13
   3359: 'Carrier 52 Power unit: Ground fault', class No Acknowledgement, trigger "DB302_HMI_Faults_Carrier52_Faults_1" bit 14
   3360: 'Spare_Fault_3360', class No Acknowledgement, trigger "DB302_HMI_Faults_Carrier52_Faults_1" bit 15
   3361: 'Carrier 52 Motion Off Fault', class No Acknowledgement, trigger "DB302_HMI_Faults_Carrier52_Faults_2" bit 0
   3362: 'Carrier 52 Motion On Fault', class No Acknowledgement, trigger "DB302_HMI_Faults_Carrier52_Faults_2" bit 1
   3363: 'Carrier 52 Spacing Fault', class No Acknowledgement, trigger "DB302_HMI_Faults_Carrier52_Faults_2" bit 2
   3364: 'Carrier 52 Duplicate Carrier Number Fault', class No Acknowledgement, trigger "DB302_HMI_Faults_Carrier52_Faults_2" bit 3
   3365: 'Spare_Fault_3365', class No Acknowledgement, trigger "DB302_HMI_Faults_Carrier52_Faults_2" bit 4
   3366: 'Spare_Fault_3366', class No Acknowledgement, trigger "DB302_HMI_Faults_Carrier52_Faults_2" bit 5
   3367: 'Spare_Fault_3367', class No Acknowledgement, trigger "DB302_HMI_Faults_Carrier52_Faults_2" bit 6
   3368: 'Spare_Fault_3368', class No Acknowledgement, trigger "DB302_HMI_Faults_Carrier52_Faults_2" bit 7
   3369: 'Spare_Fault_3369', class No Acknowledgement, trigger "DB302_HMI_Faults_Carrier52_Faults_2" bit 8
   3370: 'Spare_Fault_3370', class No Acknowledgement, trigger "DB302_HMI_Faults_Carrier52_Faults_2" bit 9
   3371: 'Spare_Fault_3371', class No Acknowledgement, trigger "DB302_HMI_Faults_Carrier52_Faults_2" bit 10
   3372: 'Spare_Fault_3372', class No Acknowledgement, trigger "DB302_HMI_Faults_Carrier52_Faults_2" bit 11
   3373: 'Spare_Fault_3373', class No Acknowledgement, trigger "DB302_HMI_Faults_Carrier52_Faults_2" bit 12
   3374: 'Spare_Fault_3374', class No Acknowledgement, trigger "DB302_HMI_Faults_Carrier52_Faults_2" bit 13
   3375: 'Spare_Fault_3375', class No Acknowledgement, trigger "DB302_HMI_Faults_Carrier52_Faults_2" bit 14
   3376: 'Spare_Fault_3376', class No Acknowledgement, trigger "DB302_HMI_Faults_Carrier52_Faults_2" bit 15
   3377: 'Spare_Fault_3377', class No Acknowledgement, trigger "DB302_HMI_Faults_Carrier52_Faults_3" bit 0
   3378: 'Spare_Fault_3378', class No Acknowledgement, trigger "DB302_HMI_Faults_Carrier52_Faults_3" bit 1
   3379: 'Spare_Fault_3379', class No Acknowledgement, trigger "DB302_HMI_Faults_Carrier52_Faults_3" bit 2
   3380: 'Spare_Fault_3380', class No Acknowledgement, trigger "DB302_HMI_Faults_Carrier52_Faults_3" bit 3
   3381: 'Spare_Fault_3381', class No Acknowledgement, trigger "DB302_HMI_Faults_Carrier52_Faults_3" bit 4
   3382: 'Spare_Fault_3382', class No Acknowledgement, trigger "DB302_HMI_Faults_Carrier52_Faults_3" bit 5
   3383: 'Spare_Fault_3383', class No Acknowledgement, trigger "DB302_HMI_Faults_Carrier52_Faults_3" bit 6
   3384: 'Spare_Fault_3384', class No Acknowledgement, trigger "DB302_HMI_Faults_Carrier52_Faults_3" bit 7
   3385: 'Spare_Fault_3385', class No Acknowledgement, trigger "DB302_HMI_Faults_Carrier52_Faults_3" bit 8
   3386: 'Spare_Fault_3386', class No Acknowledgement, trigger "DB302_HMI_Faults_Carrier52_Faults_3" bit 9
   3387: 'Spare_Fault_3387', class No Acknowledgement, trigger "DB302_HMI_Faults_Carrier52_Faults_3" bit 10
   3388: 'Spare_Fault_3388', class No Acknowledgement, trigger "DB302_HMI_Faults_Carrier52_Faults_3" bit 11
   3389: 'Spare_Fault_3389', class No Acknowledgement, trigger "DB302_HMI_Faults_Carrier52_Faults_3" bit 12
   3390: 'Spare_Fault_3390', class No Acknowledgement, trigger "DB302_HMI_Faults_Carrier52_Faults_3" bit 13
   3391: 'Spare_Fault_3391', class No Acknowledgement, trigger "DB302_HMI_Faults_Carrier52_Faults_3" bit 14
   3392: 'Spare_Fault_3392', class No Acknowledgement, trigger "DB302_HMI_Faults_Carrier52_Faults_3" bit 15
   3393: 'Carrier 53 Disconnect Open Power Fault DI11.0', class No Acknowledgement, trigger "DB302_HMI_Faults_Carrier53_Faults_0" bit 0
   3394: 'Carrier 53 Drive Profinet Comm Fault', class No Acknowledgement, trigger "DB302_HMI_Faults_Carrier53_Faults_0" bit 1
   3395: 'Carrier 53 Production Stop Not Reset', class No Acknowledgement, trigger "DB302_HMI_Faults_Carrier53_Faults_0" bit 2
